   stn[9].wipBtn[48,0] := 0;
   stn[9].wipBtn[48,1] := 0;
   stn[9].wipBtn[48,2] := 0;
   stn[9].wipBtn[48,3] := 0;
   stn[9].wipBtn[48,4] := 0;
   stn[9].wipBtn[48,5] := 0;
   stn[9].wipBtn[48,6] := 0;
   stn[9].wipBtn[48,7] := 0;
   stn[9].wipBtn[49,0] := 0;
   stn[9].wipBtn[49,1] := 0;
   stn[9].wipBtn[49,2] := 0;
   stn[9].wipBtn[49,3] := 0;
   stn[9].wipBtn[49,4] := 0;
   stn[9].wipBtn[49,5] := 0;
   stn[9].wipBtn[49,6] := 0;
   stn[9].wipBtn[49,7] := 0;
   stn[10].wipBtn[0,0] := 0;
   stn[10].wipBtn[0,1] := 0;
   stn[10].wipBtn[0,2] := 0;
   stn[10].wipBtn[0,3] := 170;
   stn[10].wipBtn[0,4] := 0;
   stn[10].wipBtn[0,5] := 0;
   stn[10].wipBtn[1,0] := 0;
   stn[10].wipBtn[1,1] := 0;
   stn[10].wipBtn[1,2] := 0;
   stn[10].wipBtn[1,3] := 0;
   stn[10].wipBtn[1,4] := 0;
   stn[10].wipBtn[1,5] := 0;
   stn[10].wipBtn[1,6] := 0;
   stn[10].wipBtn[1,7] := 0;
   stn[10].wipBtn[2,0] := 0;
   stn[10].wipBtn[2,1] := 0;
   stn[10].wipBtn[2,2] := 0;
   stn[10].wipBtn[2,3] := 0;
   stn[10].wipBtn[2,4] := 0;
   stn[10].wipBtn[2,5] := 0;
   stn[10].wipBtn[2,6] := 0;
   stn[10].wipBtn[2,7] := 0;
   stn[10].wipBtn[3,0] := 0;
   stn[10].wipBtn[3,1] := 0;
   stn[10].wipBtn[3,2] := 0;
   stn[10].wipBtn[3,3] := 0;
   stn[10].wipBtn[3,4] := 0;
   stn[10].wipBtn[3,5] := 0;
   stn[10].wipBtn[3,6] := 0;
   stn[10].wipBtn[3,7] := 0;
   stn[10].wipBtn[4,0] := 0;
   stn[10].wipBtn[4,1] := 0;
   stn[10].wipBtn[4,2] := 0;
   stn[10].wipBtn[4,3] := 0;
   stn[10].wipBtn[4,4] := 0;
   stn[10].wipBtn[4,5] := 0;
   stn[10].wipBtn[4,6] := 0;
   stn[10].wipBtn[4,7] := 0;
   stn[10].wipBtn[5,0] := 0;
   stn[10].wipBtn[5,1] := 0;
   stn[10].wipBtn[5,2] := 0;
   stn[10].wipBtn[5,3] := 0;
   stn[10].wipBtn[5,4] := 0;
   stn[10].wipBtn[5,5] := 0;
   stn[10].wipBtn[5,6] := 0;
   stn[10].wipBtn[5,7] := 0;
   stn[10].wipBtn[6,0] := 0;
   stn[10].wipBtn[6,1] := 0;
   stn[10].wipBtn[6,2] := 0;
   stn[10].wipBtn[6,3] := 0;
   stn[10].wipBtn[6,4] := 0;
   stn[10].wipBtn[6,5] := 0;
   stn[10].wipBtn[6,6] := 0;
   stn[10].wipBtn[6,7] := 0;
   stn[10].wipBtn[7,0] := 0;
   stn[10].wipBtn[7,1] := 0;
   stn[10].wipBtn[7,2] := 0;
   stn[10].wipBtn[7,3] := 0;
   stn[10].wipBtn[7,4] := 0;
   stn[10].wipBtn[7,5] := 0;
   stn[10].wipBtn[7,6] := 0;
   stn[10].wipBtn[7,7] := 0;
   stn[10].wipBtn[8,0] := 0;
   stn[10].wipBtn[8,1] := 0;
   stn[10].wipBtn[8,2] := 0;
   stn[10].wipBtn[8,3] := 0;
   stn[10].wipBtn[8,4] := 0;
   stn[10].wipBtn[8,5] := 0;
   stn[10].wipBtn[8,6] := 0;
   stn[10].wipBtn[8,7] := 0;
   stn[10].wipBtn[9,0] := 0;
   stn[10].wipBtn[9,1] := 0;
   stn[10].wipBtn[9,2] := 0;
   stn[10].wipBtn[9,3] := 0;
   stn[10].wipBtn[9,4] := 0;
   stn[10].wipBtn[9,5] := 0;
   stn[10].wipBtn[9,6] := 0;
   stn[10].wipBtn[9,7] := 0;
   stn[10].wipBtn[10,0] := 0;
   stn[10].wipBtn[10,1] := 0;
   stn[10].wipBtn[10,2] := 0;
   stn[10].wipBtn[10,3] := 0;
   stn[10].wipBtn[10,4] := 0;
   stn[10].wipBtn[10,5] := 0;
   stn[10].wipBtn[10,6] := 0;
   stn[10].wipBtn[10,7] := 0;
   stn[10].wipBtn[11,0] := 0;
   stn[10].wipBtn[11,1] := 0;
   stn[10].wipBtn[11,2] := 0;
   stn[10].wipBtn[11,3] := 0;
   stn[10].wipBtn[11,4] := 0;
   stn[10].wipBtn[11,5] := 0;
   stn[10].wipBtn[11,6] := 0;
   stn[10].wipBtn[11,7] := 0;
   stn[10].wipBtn[12,0] := 0;
   stn[10].wipBtn[12,1] := 0;
   stn[10].wipBtn[12,2] := 0;
   stn[10].wipBtn[12,3] := 0;
   stn[10].wipBtn[12,4] := 0;
   stn[10].wipBtn[12,5] := 0;
   stn[10].wipBtn[12,6] := 0;
   stn[10].wipBtn[12,7] := 0;
   stn[10].wipBtn[13,0] := 0;
   stn[10].wipBtn[13,1] := 0;
   stn[10].wipBtn[13,2] := 0;
   stn[10].wipBtn[13,3] := 0;
   stn[10].wipBtn[13,4] := 0;
   stn[10].wipBtn[13,5] := 0;
   stn[10].wipBtn[13,6] := 0;
   stn[10].wipBtn[13,7] := 0;
   stn[10].wipBtn[14,0] := 0;
   stn[10].wipBtn[14,1] := 0;
   stn[10].wipBtn[14,2] := 0;
   stn[10].wipBtn[14,3] := 0;
   stn[10].wipBtn[14,4] := 0;
   stn[10].wipBtn[14,5] := 0;
   stn[10].wipBtn[14,6] := 0;
   stn[10].wipBtn[14,7] := 0;
   stn[10].wipBtn[15,0] := 0;
   stn[10].wipBtn[15,1] := 0;
   stn[10].wipBtn[15,2] := 0;
   stn[10].wipBtn[15,3] := 0;
   stn[10].wipBtn[15,4] := 0;
   stn[10].wipBtn[15,5] := 0;
   stn[10].wipBtn[15,6] := 0;
   stn[10].wipBtn[15,7] := 0;
   stn[10].wipBtn[16,0] := 0;
   stn[10].wipBtn[16,1] := 0;
   stn[10].wipBtn[16,2] := 0;
   stn[10].wipBtn[16,3] := 0;
   stn[10].wipBtn[16,4] := 0;
   stn[10].wipBtn[16,5] := 0;
   stn[10].wipBtn[16,6] := 0;
   stn[10].wipBtn[16,7] := 0;
   stn[10].wipBtn[17,0] := 0;
   stn[10].wipBtn[17,1] := 0;
   stn[10].wipBtn[17,2] := 0;
   stn[10].wipBtn[17,3] := 0;
   stn[10].wipBtn[17,4] := 0;
   stn[10].wipBtn[17,5] := 0;
   stn[10].wipBtn[17,6] := 0;
   stn[10].wipBtn[17,7] := 0;
   stn[10].wipBtn[18,0] := 0;
   stn[10].wipBtn[18,1] := 0;
   stn[10].wipBtn[18,2] := 0;
   stn[10].wipBtn[18,3] := 0;
   stn[10].wipBtn[18,4] := 0;
   stn[10].wipBtn[18,5] := 0;
   stn[10].wipBtn[18,6] := 0;
   stn[10].wipBtn[18,7] := 0;
   stn[10].wipBtn[19,0] := 0;
   stn[10].wipBtn[19,1] := 0;
   stn[10].wipBtn[19,2] := 0;
   stn[10].wipBtn[19,3] := 0;
   stn[10].wipBtn[19,4] := 0;
   stn[10].wipBtn[19,5] := 0;
   stn[10].wipBtn[19,6] := 0;
   stn[10].wipBtn[19,7] := 0;
   stn[10].wipBtn[20,0] := 0;
   stn[10].wipBtn[20,1] := 0;
   stn[10].wipBtn[20,2] := 0;
   stn[10].wipBtn[20,3] := 0;
   stn[10].wipBtn[20,4] := 0;
   stn[10].wipBtn[20,5] := 0;
   stn[10].wipBtn[20,6] := 0;
   stn[10].wipBtn[20,7] := 0;
   stn[10].wipBtn[21,0] := 0;
   stn[10].wipBtn[21,1] := 0;
   stn[10].wipBtn[21,2] := 0;
   stn[10].wipBtn[21,3] := 0;
   stn[10].wipBtn[21,4] := 0;
   stn[10].wipBtn[21,5] := 0;
   stn[10].wipBtn[21,6] := 0;
   stn[10].wipBtn[21,7] := 0;
   stn[10].wipBtn[22,0] := 0;
   stn[10].wipBtn[22,1] := 0;
   stn[10].wipBtn[22,2] := 0;
   stn[10].wipBtn[22,3] := 0;
   stn[10].wipBtn[22,4] := 0;
   stn[10].wipBtn[22,5] := 0;
   stn[10].wipBtn[22,6] := 0;
   stn[10].wipBtn[22,7] := 0;
   stn[10].wipBtn[23,0] := 0;
   stn[10].wipBtn[23,1] := 0;
   stn[10].wipBtn[23,2] := 0;
   stn[10].wipBtn[23,3] := 0;
   stn[10].wipBtn[23,4] := 0;
   stn[10].wipBtn[23,5] := 0;
   stn[10].wipBtn[23,6] := 0;
   stn[10].wipBtn[23,7] := 0;
   stn[10].wipBtn[24,0] := 0;
   stn[10].wipBtn[24,1] := 0;
   stn[10].wipBtn[24,2] := 0;
   stn[10].wipBtn[24,3] := 0;
   stn[10].wipBtn[24,4] := 0;
   stn[10].wipBtn[24,5] := 0;
   stn[10].wipBtn[24,6] := 0;
   stn[10].wipBtn[24,7] := 0;
   stn[10].wipBtn[25,0] := 0;
   stn[10].wipBtn[25,1] := 0;
   stn[10].wipBtn[25,2] := 0;
   stn[10].wipBtn[25,3] := 0;
   stn[10].wipBtn[25,4] := 0;
   stn[10].wipBtn[25,5] := 0;
   stn[10].wipBtn[25,6] := 0;
   stn[10].wipBtn[25,7] := 0;
   stn[10].wipBtn[26,0] := 0;
   stn[10].wipBtn[26,1] := 0;
   stn[10].wipBtn[26,2] := 0;
   stn[10].wipBtn[26,3] := 0;
   stn[10].wipBtn[26,4] := 0;
   stn[10].wipBtn[26,5] := 0;
   stn[10].wipBtn[26,6] := 0;
   stn[10].wipBtn[26,7] := 0;
   stn[10].wipBtn[27,0] := 0;
   stn[10].wipBtn[27,1] := 0;
   stn[10].wipBtn[27,2] := 0;
   stn[10].wipBtn[27,3] := 0;
   stn[10].wipBtn[27,4] := 0;
   stn[10].wipBtn[27,5] := 0;
   stn[10].wipBtn[27,6] := 0;
   stn[10].wipBtn[27,7] := 0;
   stn[10].wipBtn[28,0] := 0;
   stn[10].wipBtn[28,1] := 0;
   stn[10].wipBtn[28,2] := 0;
   stn[10].wipBtn[28,3] := 0;
   stn[10].wipBtn[28,4] := 0;
   stn[10].wipBtn[28,5] := 0;
   stn[10].wipBtn[28,6] := 0;
   stn[10].wipBtn[28,7] := 0;
   stn[10].wipBtn[29,0] := 0;
   stn[10].wipBtn[29,1] := 0;
   stn[10].wipBtn[29,2] := 0;
   stn[10].wipBtn[29,3] := 0;
   stn[10].wipBtn[29,4] := 0;
   stn[10].wipBtn[29,5] := 0;
   stn[10].wipBtn[29,6] := 0;
   stn[10].wipBtn[29,7] := 0;
   stn[10].wipBtn[30,0] := 0;
   stn[10].wipBtn[30,1] := 0;
   stn[10].wipBtn[30,2] := 0;
   stn[10].wipBtn[30,3] := 0;
   stn[10].wipBtn[30,4] := 0;
   stn[10].wipBtn[30,5] := 0;
   stn[10].wipBtn[30,6] := 0;
   stn[10].wipBtn[30,7] := 0;
   stn[10].wipBtn[31,0] := 0;
   stn[10].wipBtn[31,1] := 0;
   stn[10].wipBtn[31,2] := 0;
   stn[10].wipBtn[31,3] := 0;
   stn[10].wipBtn[31,4] := 0;
   stn[10].wipBtn[31,5] := 0;
   stn[10].wipBtn[31,6] := 0;
   stn[10].wipBtn[31,7] := 0;
   stn[10].wipBtn[32,0] := 0;
   stn[10].wipBtn[32,1] := 0;
   stn[10].wipBtn[32,2] := 0;
   stn[10].wipBtn[32,3] := 0;
   stn[10].wipBtn[32,4] := 0;
   stn[10].wipBtn[32,5] := 0;
   stn[10].wipBtn[32,6] := 0;
   stn[10].wipBtn[32,7] := 0;
   stn[10].wipBtn[33,0] := 0;
   stn[10].wipBtn[33,1] := 0;
   stn[10].wipBtn[33,2] := 0;
   stn[10].wipBtn[33,3] := 0;
   stn[10].wipBtn[33,4] := 0;
   stn[10].wipBtn[33,5] := 0;
   stn[10].wipBtn[33,6] := 0;
   stn[10].wipBtn[33,7] := 0;
   stn[10].wipBtn[34,0] := 0;
   stn[10].wipBtn[34,1] := 0;
   stn[10].wipBtn[34,2] := 0;
   stn[10].wipBtn[34,3] := 0;
   stn[10].wipBtn[34,4] := 0;
   stn[10].wipBtn[34,5] := 0;
   stn[10].wipBtn[34,6] := 0;
   stn[10].wipBtn[34,7] := 0;
   stn[10].wipBtn[35,0] := 0;
   stn[10].wipBtn[35,1] := 0;
   stn[10].wipBtn[35,2] := 0;
   stn[10].wipBtn[35,3] := 0;
   stn[10].wipBtn[35,4] := 0;
   stn[10].wipBtn[35,5] := 0;
   stn[10].wipBtn[35,6] := 0;
   stn[10].wipBtn[35,7] := 0;
   stn[10].wipBtn[36,0] := 0;
   stn[10].wipBtn[36,1] := 0;
   stn[10].wipBtn[36,2] := 0;
   stn[10].wipBtn[36,3] := 0;
   stn[10].wipBtn[36,4] := 0;
   stn[10].wipBtn[36,5] := 0;
   stn[10].wipBtn[36,6] := 0;
   stn[10].wipBtn[36,7] := 0;
   stn[10].wipBtn[37,0] := 0;
   stn[10].wipBtn[37,1] := 0;
   stn[10].wipBtn[37,2] := 0;
   stn[10].wipBtn[37,3] := 0;
   stn[10].wipBtn[37,4] := 0;
   stn[10].wipBtn[37,5] := 0;
   stn[10].wipBtn[37,6] := 0;
   stn[10].wipBtn[37,7] := 0;
   stn[10].wipBtn[38,0] := 0;
   stn[10].wipBtn[38,1] := 0;
   stn[10].wipBtn[38,2] := 0;
   stn[10].wipBtn[38,3] := 0;
   stn[10].wipBtn[38,4] := 0;
   stn[10].wipBtn[38,5] := 0;
   stn[10].wipBtn[38,6] := 0;
   stn[10].wipBtn[38,7] := 0;
   stn[10].wipBtn[39,0] := 0;
   stn[10].wipBtn[39,1] := 0;
   stn[10].wipBtn[39,2] := 0;
   stn[10].wipBtn[39,3] := 0;
   stn[10].wipBtn[39,4] := 0;
   stn[10].wipBtn[39,5] := 0;
   stn[10].wipBtn[39,6] := 0;
   stn[10].wipBtn[39,7] := 0;
   stn[10].wipBtn[40,0] := 0;
   stn[10].wipBtn[40,1] := 0;
   stn[10].wipBtn[40,2] := 0;
   stn[10].wipBtn[40,3] := 0;
   stn[10].wipBtn[40,4] := 0;
   stn[10].wipBtn[40,5] := 0;
   stn[10].wipBtn[40,6] := 0;
   stn[10].wipBtn[40,7] := 0;
   stn[10].wipBtn[41,0] := 0;
   stn[10].wipBtn[41,1] := 0;
   stn[10].wipBtn[41,2] := 0;
   stn[10].wipBtn[41,3] := 0;
   stn[10].wipBtn[41,4] := 0;
   stn[10].wipBtn[41,5] := 0;
   stn[10].wipBtn[41,6] := 0;
   stn[10].wipBtn[41,7] := 0;
   stn[10].wipBtn[42,0] := 0;
   stn[10].wipBtn[42,1] := 0;
   stn[10].wipBtn[42,2] := 0;
   stn[10].wipBtn[42,3] := 0;
   stn[10].wipBtn[42,4] := 0;
   stn[10].wipBtn[42,5] := 0;
   stn[10].wipBtn[42,6] := 0;
   stn[10].wipBtn[42,7] := 0;
   stn[10].wipBtn[43,0] := 0;
   stn[10].wipBtn[43,1] := 0;
   stn[10].wipBtn[43,2] := 0;
   stn[10].wipBtn[43,3] := 0;
   stn[10].wipBtn[43,4] := 0;
   stn[10].wipBtn[43,5] := 0;
   stn[10].wipBtn[43,6] := 0;
   stn[10].wipBtn[43,7] := 0;
   stn[10].wipBtn[44,0] := 0;
   stn[10].wipBtn[44,1] := 0;
   stn[10].wipBtn[44,2] := 0;
   stn[10].wipBtn[44,3] := 0;
   stn[10].wipBtn[44,4] := 0;
   stn[10].wipBtn[44,5] := 0;
   stn[10].wipBtn[44,6] := 0;
   stn[10].wipBtn[44,7] := 0;
   stn[10].wipBtn[45,0] := 0;
   stn[10].wipBtn[45,1] := 0;
   stn[10].wipBtn[45,2] := 0;
   stn[10].wipBtn[45,3] := 0;
   stn[10].wipBtn[45,4] := 0;
   stn[10].wipBtn[45,5] := 0;
   stn[10].wipBtn[45,6] := 0;
   stn[10].wipBtn[45,7] := 0;
   stn[10].wipBtn[46,0] := 0;
   stn[10].wipBtn[46,1] := 0;
   stn[10].wipBtn[46,2] := 0;
   stn[10].wipBtn[46,3] := 0;
   stn[10].wipBtn[46,4] := 0;
   stn[10].wipBtn[46,5] := 0;
   stn[10].wipBtn[46,6] := 0;
   stn[10].wipBtn[46,7] := 0;
   stn[10].wipBtn[47,0] := 0;
   stn[10].wipBtn[47,1] := 0;
   stn[10].wipBtn[47,2] := 0;
   stn[10].wipBtn[47,3] := 0;
   stn[10].wipBtn[47,4] := 0;
   stn[10].wipBtn[47,5] := 0;
   stn[10].wipBtn[47,6] := 0;
   stn[10].wipBtn[47,7] := 0;
   stn[10].wipBtn[48,0] := 0;
   stn[10].wipBtn[48,1] := 0;
   stn[10].wipBtn[48,2] := 0;
   stn[10].wipBtn[48,3] := 0;
   stn[10].wipBtn[48,4] := 0;
   stn[10].wipBtn[48,5] := 0;
   stn[10].wipBtn[48,6] := 0;
   stn[10].wipBtn[48,7] := 0;
   stn[10].wipBtn[49,0] := 0;
   stn[10].wipBtn[49,1] := 0;
   stn[10].wipBtn[49,2] := 0;
   stn[10].wipBtn[49,3] := 0;
   stn[10].wipBtn[49,4] := 0;
   stn[10].wipBtn[49,5] := 0;
   stn[10].wipBtn[49,6] := 0;
   stn[10].wipBtn[49,7] := 0;
   stn[11].wipBtn[0,0] := 0;
   stn[11].wipBtn[0,1] := 0;
   stn[11].wipBtn[0,2] := 0;
   stn[11].wipBtn[0,4] := 0;
   stn[11].wipBtn[0,5] := 0;
   stn[11].wipBtn[0,7] := 20;
   stn[11].wipBtn[1,0] := 0;
   stn[11].wipBtn[1,1] := 0;
   stn[11].wipBtn[1,2] := 0;
   stn[11].wipBtn[1,3] := 0;
   stn[11].wipBtn[1,4] := 0;
   stn[11].wipBtn[1,5] := 0;
   stn[11].wipBtn[1,6] := 0;
   stn[11].wipBtn[1,7] := 0;
   stn[11].wipBtn[2,0] := 0;
   stn[11].wipBtn[2,1] := 0;
   stn[11].wipBtn[2,2] := 0;
   stn[11].wipBtn[2,3] := 0;
   stn[11].wipBtn[2,4] := 0;
   stn[11].wipBtn[2,5] := 0;
   stn[11].wipBtn[2,6] := 0;
   stn[11].wipBtn[2,7] := 0;
   stn[11].wipBtn[3,0] := 0;
   stn[11].wipBtn[3,1] := 0;
   stn[11].wipBtn[3,2] := 0;
   stn[11].wipBtn[3,3] := 0;
   stn[11].wipBtn[3,4] := 0;
   stn[11].wipBtn[3,5] := 0;
   stn[11].wipBtn[3,6] := 0;
   stn[11].wipBtn[3,7] := 0;
   stn[11].wipBtn[4,0] := 0;
   stn[11].wipBtn[4,1] := 0;
   stn[11].wipBtn[4,2] := 0;
   stn[11].wipBtn[4,3] := 0;
   stn[11].wipBtn[4,4] := 0;
   stn[11].wipBtn[4,5] := 0;
   stn[11].wipBtn[4,6] := 0;
   stn[11].wipBtn[4,7] := 0;
   stn[11].wipBtn[5,0] := 0;
   stn[11].wipBtn[5,1] := 0;
   stn[11].wipBtn[5,2] := 0;
   stn[11].wipBtn[5,3] := 0;
   stn[11].wipBtn[5,4] := 0;
   stn[11].wipBtn[5,5] := 0;
   stn[11].wipBtn[5,6] := 0;
   stn[11].wipBtn[5,7] := 0;
   stn[11].wipBtn[6,0] := 0;
   stn[11].wipBtn[6,1] := 0;
   stn[11].wipBtn[6,2] := 0;
   stn[11].wipBtn[6,3] := 0;
   stn[11].wipBtn[6,4] := 0;
   stn[11].wipBtn[6,5] := 0;
   stn[11].wipBtn[6,6] := 0;
   stn[11].wipBtn[6,7] := 0;
   stn[11].wipBtn[7,0] := 0;
   stn[11].wipBtn[7,1] := 0;
   stn[11].wipBtn[7,2] := 0;
   stn[11].wipBtn[7,3] := 0;
   stn[11].wipBtn[7,4] := 0;
   stn[11].wipBtn[7,5] := 0;
   stn[11].wipBtn[7,6] := 0;
   stn[11].wipBtn[7,7] := 0;
   stn[11].wipBtn[8,0] := 0;
   stn[11].wipBtn[8,1] := 0;
   stn[11].wipBtn[8,2] := 0;
   stn[11].wipBtn[8,3] := 0;
   stn[11].wipBtn[8,4] := 0;
   stn[11].wipBtn[8,5] := 0;
   stn[11].wipBtn[8,6] := 0;
   stn[11].wipBtn[8,7] := 0;
   stn[11].wipBtn[9,0] := 0;
   stn[11].wipBtn[9,1] := 0;
   stn[11].wipBtn[9,2] := 0;
   stn[11].wipBtn[9,3] := 0;
   stn[11].wipBtn[9,4] := 0;
   stn[11].wipBtn[9,5] := 0;
   stn[11].wipBtn[9,6] := 0;
   stn[11].wipBtn[9,7] := 0;
   stn[11].wipBtn[10,0] := 0;
   stn[11].wipBtn[10,1] := 0;
   stn[11].wipBtn[10,2] := 0;
   stn[11].wipBtn[10,3] := 0;
   stn[11].wipBtn[10,4] := 0;
   stn[11].wipBtn[10,5] := 0;
   stn[11].wipBtn[10,6] := 0;
   stn[11].wipBtn[10,7] := 0;
   stn[11].wipBtn[11,0] := 0;
   stn[11].wipBtn[11,1] := 0;
   stn[11].wipBtn[11,2] := 0;
   stn[11].wipBtn[11,3] := 0;
   stn[11].wipBtn[11,4] := 0;
   stn[11].wipBtn[11,5] := 0;
   stn[11].wipBtn[11,6] := 0;
   stn[11].wipBtn[11,7] := 0;
   stn[11].wipBtn[12,0] := 0;
   stn[11].wipBtn[12,1] := 0;
   stn[11].wipBtn[12,2] := 0;
   stn[11].wipBtn[12,3] := 0;
   stn[11].wipBtn[12,4] := 0;
   stn[11].wipBtn[12,5] := 0;
   stn[11].wipBtn[12,6] := 0;
   stn[11].wipBtn[12,7] := 0;
   stn[11].wipBtn[13,0] := 0;
   stn[11].wipBtn[13,1] := 0;
   stn[11].wipBtn[13,2] := 0;
   stn[11].wipBtn[13,3] := 0;
   stn[11].wipBtn[13,4] := 0;
   stn[11].wipBtn[13,5] := 0;
   stn[11].wipBtn[13,6] := 0;
   stn[11].wipBtn[13,7] := 0;
   stn[11].wipBtn[14,0] := 0;
   stn[11].wipBtn[14,1] := 0;
   stn[11].wipBtn[14,2] := 0;
   stn[11].wipBtn[14,3] := 0;
   stn[11].wipBtn[14,4] := 0;
   stn[11].wipBtn[14,5] := 0;
   stn[11].wipBtn[14,6] := 0;
   stn[11].wipBtn[14,7] := 0;
   stn[11].wipBtn[15,0] := 0;
   stn[11].wipBtn[15,1] := 0;
   stn[11].wipBtn[15,2] := 0;
   stn[11].wipBtn[15,3] := 0;
   stn[11].wipBtn[15,4] := 0;
   stn[11].wipBtn[15,5] := 0;
   stn[11].wipBtn[15,6] := 0;
   stn[11].wipBtn[15,7] := 0;
   stn[11].wipBtn[16,0] := 0;
   stn[11].wipBtn[16,1] := 0;
   stn[11].wipBtn[16,2] := 0;
   stn[11].wipBtn[16,3] := 0;
   stn[11].wipBtn[16,4] := 0;
   stn[11].wipBtn[16,5] := 0;
   stn[11].wipBtn[16,6] := 0;
   stn[11].wipBtn[16,7] := 0;
   stn[11].wipBtn[17,0] := 0;
   stn[11].wipBtn[17,1] := 0;
   stn[11].wipBtn[17,2] := 0;
   stn[11].wipBtn[17,3] := 0;
   stn[11].wipBtn[17,4] := 0;
   stn[11].wipBtn[17,5] := 0;
   stn[11].wipBtn[17,6] := 0;
   stn[11].wipBtn[17,7] := 0;
   stn[11].wipBtn[18,0] := 0;
   stn[11].wipBtn[18,1] := 0;
   stn[11].wipBtn[18,2] := 0;
   stn[11].wipBtn[18,3] := 0;
   stn[11].wipBtn[18,4] := 0;
   stn[11].wipBtn[18,5] := 0;
   stn[11].wipBtn[18,6] := 0;
   stn[11].wipBtn[18,7] := 0;
   stn[11].wipBtn[19,0] := 0;
   stn[11].wipBtn[19,1] := 0;
   stn[11].wipBtn[19,2] := 0;
   stn[11].wipBtn[19,3] := 0;
   stn[11].wipBtn[19,4] := 0;
   stn[11].wipBtn[19,5] := 0;
   stn[11].wipBtn[19,6] := 0;
   stn[11].wipBtn[19,7] := 0;
   stn[11].wipBtn[20,0] := 0;
   stn[11].wipBtn[20,1] := 0;
   stn[11].wipBtn[20,2] := 0;
   stn[11].wipBtn[20,3] := 0;
   stn[11].wipBtn[20,4] := 0;
   stn[11].wipBtn[20,5] := 0;
   stn[11].wipBtn[20,6] := 0;
   stn[11].wipBtn[20,7] := 0;
   stn[11].wipBtn[21,0] := 0;
   stn[11].wipBtn[21,1] := 0;
   stn[11].wipBtn[21,2] := 0;
   stn[11].wipBtn[21,3] := 0;
   stn[11].wipBtn[21,4] := 0;
   stn[11].wipBtn[21,5] := 0;
   stn[11].wipBtn[21,6] := 0;
   stn[11].wipBtn[21,7] := 0;
   stn[11].wipBtn[22,0] := 0;
   stn[11].wipBtn[22,1] := 0;
   stn[11].wipBtn[22,2] := 0;
   stn[11].wipBtn[22,3] := 0;
   stn[11].wipBtn[22,4] := 0;
   stn[11].wipBtn[22,5] := 0;
   stn[11].wipBtn[22,6] := 0;
   stn[11].wipBtn[22,7] := 0;
   stn[11].wipBtn[23,0] := 0;
   stn[11].wipBtn[23,1] := 0;
   stn[11].wipBtn[23,2] := 0;
   stn[11].wipBtn[23,3] := 0;
   stn[11].wipBtn[23,4] := 0;
   stn[11].wipBtn[23,5] := 0;
   stn[11].wipBtn[23,6] := 0;
   stn[11].wipBtn[23,7] := 0;
   stn[11].wipBtn[24,0] := 0;
   stn[11].wipBtn[24,1] := 0;
   stn[11].wipBtn[24,2] := 0;
   stn[11].wipBtn[24,3] := 0;
   stn[11].wipBtn[24,4] := 0;
   stn[11].wipBtn[24,5] := 0;
   stn[11].wipBtn[24,6] := 0;
   stn[11].wipBtn[24,7] := 0;
   stn[11].wipBtn[25,0] := 0;
   stn[11].wipBtn[25,1] := 0;
   stn[11].wipBtn[25,2] := 0;
   stn[11].wipBtn[25,3] := 0;
   stn[11].wipBtn[25,4] := 0;
   stn[11].wipBtn[25,5] := 0;
   stn[11].wipBtn[25,6] := 0;
   stn[11].wipBtn[25,7] := 0;
   stn[11].wipBtn[26,0] := 0;
   stn[11].wipBtn[26,1] := 0;
   stn[11].wipBtn[26,2] := 0;
   stn[11].wipBtn[26,3] := 0;
   stn[11].wipBtn[26,4] := 0;
   stn[11].wipBtn[26,5] := 0;
   stn[11].wipBtn[26,6] := 0;
   stn[11].wipBtn[26,7] := 0;
   stn[11].wipBtn[27,0] := 0;
   stn[11].wipBtn[27,1] := 0;
   stn[11].wipBtn[27,2] := 0;
   stn[11].wipBtn[27,3] := 0;
   stn[11].wipBtn[27,4] := 0;
   stn[11].wipBtn[27,5] := 0;
   stn[11].wipBtn[27,6] := 0;
   stn[11].wipBtn[27,7] := 0;
   stn[11].wipBtn[28,0] := 0;
   stn[11].wipBtn[28,1] := 0;
   stn[11].wipBtn[28,2] := 0;
   stn[11].wipBtn[28,3] := 0;
   stn[11].wipBtn[28,4] := 0;
   stn[11].wipBtn[28,5] := 0;
   stn[11].wipBtn[28,6] := 0;
   stn[11].wipBtn[28,7] := 0;
   stn[11].wipBtn[29,0] := 0;
   stn[11].wipBtn[29,1] := 0;
   stn[11].wipBtn[29,2] := 0;
   stn[11].wipBtn[29,3] := 0;
   stn[11].wipBtn[29,4] := 0;
   stn[11].wipBtn[29,5] := 0;
   stn[11].wipBtn[29,6] := 0;
   stn[11].wipBtn[29,7] := 0;
   stn[11].wipBtn[30,0] := 0;
   stn[11].wipBtn[30,1] := 0;
   stn[11].wipBtn[30,2] := 0;
   stn[11].wipBtn[30,3] := 0;
   stn[11].wipBtn[30,4] := 0;
   stn[11].wipBtn[30,5] := 0;
   stn[11].wipBtn[30,6] := 0;
   stn[11].wipBtn[30,7] := 0;
   stn[11].wipBtn[31,0] := 0;
   stn[11].wipBtn[31,1] := 0;
   stn[11].wipBtn[31,2] := 0;
   stn[11].wipBtn[31,3] := 0;
   stn[11].wipBtn[31,4] := 0;
   stn[11].wipBtn[31,5] := 0;
   stn[11].wipBtn[31,6] := 0;
   stn[11].wipBtn[31,7] := 0;
   stn[11].wipBtn[32,0] := 0;
   stn[11].wipBtn[32,1] := 0;
   stn[11].wipBtn[32,2] := 0;
   stn[11].wipBtn[32,3] := 0;
   stn[11].wipBtn[32,4] := 0;
   stn[11].wipBtn[32,5] := 0;
   stn[11].wipBtn[32,6] := 0;
   stn[11].wipBtn[32,7] := 0;
   stn[11].wipBtn[33,0] := 0;
   stn[11].wipBtn[33,1] := 0;
   stn[11].wipBtn[33,2] := 0;
   stn[11].wipBtn[33,3] := 0;
   stn[11].wipBtn[33,4] := 0;
   stn[11].wipBtn[33,5] := 0;
   stn[11].wipBtn[33,6] := 0;
   stn[11].wipBtn[33,7] := 0;
   stn[11].wipBtn[34,0] := 0;
   stn[11].wipBtn[34,1] := 0;
   stn[11].wipBtn[34,2] := 0;
   stn[11].wipBtn[34,3] := 0;
   stn[11].wipBtn[34,4] := 0;
   stn[11].wipBtn[34,5] := 0;
   stn[11].wipBtn[34,6] := 0;
   stn[11].wipBtn[34,7] := 0;
   stn[11].wipBtn[35,0] := 0;
   stn[11].wipBtn[35,1] := 0;
   stn[11].wipBtn[35,2] := 0;
   stn[11].wipBtn[35,3] := 0;
   stn[11].wipBtn[35,4] := 0;
   stn[11].wipBtn[35,5] := 0;
   stn[11].wipBtn[35,6] := 0;
   stn[11].wipBtn[35,7] := 0;
   stn[11].wipBtn[36,0] := 0;
   stn[11].wipBtn[36,1] := 0;
   stn[11].wipBtn[36,2] := 0;
   stn[11].wipBtn[36,3] := 0;
   stn[11].wipBtn[36,4] := 0;
   stn[11].wipBtn[36,5] := 0;
   stn[11].wipBtn[36,6] := 0;
   stn[11].wipBtn[36,7] := 0;
   stn[11].wipBtn[37,0] := 0;
   stn[11].wipBtn[37,1] := 0;
   stn[11].wipBtn[37,2] := 0;
   stn[11].wipBtn[37,3] := 0;
   stn[11].wipBtn[37,4] := 0;
   stn[11].wipBtn[37,5] := 0;
   stn[11].wipBtn[37,6] := 0;
   stn[11].wipBtn[37,7] := 0;
   stn[11].wipBtn[38,0] := 0;
   stn[11].wipBtn[38,1] := 0;
   stn[11].wipBtn[38,2] := 0;
   stn[11].wipBtn[38,3] := 0;
   stn[11].wipBtn[38,4] := 0;
   stn[11].wipBtn[38,5] := 0;
   stn[11].wipBtn[38,6] := 0;
   stn[11].wipBtn[38,7] := 0;
   stn[11].wipBtn[39,0] := 0;
   stn[11].wipBtn[39,1] := 0;
   stn[11].wipBtn[39,2] := 0;
   stn[11].wipBtn[39,3] := 0;
   stn[11].wipBtn[39,4] := 0;
   stn[11].wipBtn[39,5] := 0;
   stn[11].wipBtn[39,6] := 0;
   stn[11].wipBtn[39,7] := 0;
   stn[11].wipBtn[40,0] := 0;
   stn[11].wipBtn[40,1] := 0;
   stn[11].wipBtn[40,2] := 0;
   stn[11].wipBtn[40,3] := 0;
   stn[11].wipBtn[40,4] := 0;
   stn[11].wipBtn[40,5] := 0;
   stn[11].wipBtn[40,6] := 0;
   stn[11].wipBtn[40,7] := 0;
   stn[11].wipBtn[41,0] := 0;
   stn[11].wipBtn[41,1] := 0;
   stn[11].wipBtn[41,2] := 0;
   stn[11].wipBtn[41,3] := 0;
   stn[11].wipBtn[41,4] := 0;
   stn[11].wipBtn[41,5] := 0;
   stn[11].wipBtn[41,6] := 0;
   stn[11].wipBtn[41,7] := 0;
   stn[11].wipBtn[42,0] := 0;
   stn[11].wipBtn[42,1] := 0;
   stn[11].wipBtn[42,2] := 0;
   stn[11].wipBtn[42,3] := 0;
   stn[11].wipBtn[42,4] := 0;
   stn[11].wipBtn[42,5] := 0;
   stn[11].wipBtn[42,6] := 0;
   stn[11].wipBtn[42,7] := 0;
   stn[11].wipBtn[43,0] := 0;
   stn[11].wipBtn[43,1] := 0;
   stn[11].wipBtn[43,2] := 0;
   stn[11].wipBtn[43,3] := 0;
   stn[11].wipBtn[43,4] := 0;
   stn[11].wipBtn[43,5] := 0;
   stn[11].wipBtn[43,6] := 0;
   stn[11].wipBtn[43,7] := 0;
   stn[11].wipBtn[44,0] := 0;
   stn[11].wipBtn[44,1] := 0;
   stn[11].wipBtn[44,2] := 0;
   stn[11].wipBtn[44,3] := 0;
   stn[11].wipBtn[44,4] := 0;
   stn[11].wipBtn[44,5] := 0;
   stn[11].wipBtn[44,6] := 0;
   stn[11].wipBtn[44,7] := 0;
   stn[11].wipBtn[45,0] := 0;
   stn[11].wipBtn[45,1] := 0;
   stn[11].wipBtn[45,2] := 0;
   stn[11].wipBtn[45,3] := 0;
   stn[11].wipBtn[45,4] := 0;
   stn[11].wipBtn[45,5] := 0;
   stn[11].wipBtn[45,6] := 0;
   stn[11].wipBtn[45,7] := 0;
   stn[11].wipBtn[46,0] := 0;
   stn[11].wipBtn[46,1] := 0;
   stn[11].wipBtn[46,2] := 0;
   stn[11].wipBtn[46,3] := 0;
   stn[11].wipBtn[46,4] := 0;
   stn[11].wipBtn[46,5] := 0;
   stn[11].wipBtn[46,6] := 0;
   stn[11].wipBtn[46,7] := 0;
   stn[11].wipBtn[47,0] := 0;
   stn[11].wipBtn[47,1] := 0;
   stn[11].wipBtn[47,2] := 0;
   stn[11].wipBtn[47,3] := 0;
   stn[11].wipBtn[47,4] := 0;
   stn[11].wipBtn[47,5] := 0;
   stn[11].wipBtn[47,6] := 0;
   stn[11].wipBtn[47,7] := 0;
   stn[11].wipBtn[48,0] := 0;
   stn[11].wipBtn[48,1] := 0;
   stn[11].wipBtn[48,2] := 0;
   stn[11].wipBtn[48,3] := 0;
   stn[11].wipBtn[48,4] := 0;
   stn[11].wipBtn[48,5] := 0;
   stn[11].wipBtn[48,6] := 0;
   stn[11].wipBtn[48,7] := 0;
   stn[11].wipBtn[49,0] := 0;
   stn[11].wipBtn[49,1] := 0;
   stn[11].wipBtn[49,2] := 0;
   stn[11].wipBtn[49,3] := 0;
   stn[11].wipBtn[49,4] := 0;
   stn[11].wipBtn[49,5] := 0;
   stn[11].wipBtn[49,6] := 0;
   stn[11].wipBtn[49,7] := 0;
   stn[12].wipBtn[0,0] := 0;
   stn[12].wipBtn[0,1] := 80;
   stn[12].wipBtn[0,4] := 0;
   stn[12].wipBtn[1,0] := 0;
   stn[12].wipBtn[1,1] := 0;
   stn[12].wipBtn[1,2] := 0;
   stn[12].wipBtn[1,3] := 0;
   stn[12].wipBtn[1,4] := 0;
   stn[12].wipBtn[1,5] := 0;
   stn[12].wipBtn[1,6] := 0;
   stn[12].wipBtn[1,7] := 0;
   stn[12].wipBtn[2,0] := 0;
   stn[12].wipBtn[2,1] := 0;
   stn[12].wipBtn[2,2] := 0;
   stn[12].wipBtn[2,3] := 0;
   stn[12].wipBtn[2,4] := 0;
   stn[12].wipBtn[2,5] := 0;
   stn[12].wipBtn[2,6] := 0;
   stn[12].wipBtn[2,7] := 0;
   stn[12].wipBtn[3,0] := 0;
   stn[12].wipBtn[3,1] := 0;
   stn[12].wipBtn[3,2] := 0;
   stn[12].wipBtn[3,3] := 0;
   stn[12].wipBtn[3,4] := 0;
   stn[12].wipBtn[3,5] := 0;
   stn[12].wipBtn[3,6] := 0;
   stn[12].wipBtn[3,7] := 0;
   stn[12].wipBtn[4,0] := 0;
   stn[12].wipBtn[4,1] := 0;
   stn[12].wipBtn[4,2] := 0;
   stn[12].wipBtn[4,3] := 0;
   stn[12].wipBtn[4,4] := 0;
   stn[12].wipBtn[4,5] := 0;
   stn[12].wipBtn[4,6] := 0;
   stn[12].wipBtn[4,7] := 0;
   stn[12].wipBtn[5,0] := 0;
   stn[12].wipBtn[5,1] := 0;
   stn[12].wipBtn[5,2] := 0;
   stn[12].wipBtn[5,3] := 0;
   stn[12].wipBtn[5,4] := 0;
   stn[12].wipBtn[5,5] := 0;
   stn[12].wipBtn[5,6] := 0;
   stn[12].wipBtn[5,7] := 0;
   stn[12].wipBtn[6,0] := 0;
   stn[12].wipBtn[6,1] := 0;
   stn[12].wipBtn[6,2] := 0;
   stn[12].wipBtn[6,3] := 0;
   stn[12].wipBtn[6,4] := 0;
   stn[12].wipBtn[6,5] := 0;
   stn[12].wipBtn[6,6] := 0;
   stn[12].wipBtn[6,7] := 0;
   stn[12].wipBtn[7,0] := 0;
   stn[12].wipBtn[7,1] := 0;
   stn[12].wipBtn[7,2] := 0;
   stn[12].wipBtn[7,3] := 0;
   stn[12].wipBtn[7,4] := 0;
   stn[12].wipBtn[7,5] := 0;
   stn[12].wipBtn[7,6] := 0;
   stn[12].wipBtn[7,7] := 0;
   stn[12].wipBtn[8,0] := 0;
   stn[12].wipBtn[8,1] := 0;
   stn[12].wipBtn[8,2] := 0;
   stn[12].wipBtn[8,3] := 0;
   stn[12].wipBtn[8,4] := 0;
   stn[12].wipBtn[8,5] := 0;
   stn[12].wipBtn[8,6] := 0;
   stn[12].wipBtn[8,7] := 0;
   stn[12].wipBtn[9,0] := 0;
   stn[12].wipBtn[9,1] := 0;
   stn[12].wipBtn[9,2] := 0;
   stn[12].wipBtn[9,3] := 0;
   stn[12].wipBtn[9,4] := 0;
   stn[12].wipBtn[9,5] := 0;
   stn[12].wipBtn[9,6] := 0;
   stn[12].wipBtn[9,7] := 0;
   stn[12].wipBtn[10,0] := 0;
   stn[12].wipBtn[10,1] := 0;
   stn[12].wipBtn[10,2] := 0;
   stn[12].wipBtn[10,3] := 0;
   stn[12].wipBtn[10,4] := 0;
   stn[12].wipBtn[10,5] := 0;
   stn[12].wipBtn[10,6] := 0;
   stn[12].wipBtn[10,7] := 0;
   stn[12].wipBtn[11,0] := 0;
   stn[12].wipBtn[11,1] := 0;
   stn[12].wipBtn[11,2] := 0;
   stn[12].wipBtn[11,3] := 0;
   stn[12].wipBtn[11,4] := 0;
   stn[12].wipBtn[11,5] := 0;
   stn[12].wipBtn[11,6] := 0;
   stn[12].wipBtn[11,7] := 0;
   stn[12].wipBtn[12,0] := 0;
   stn[12].wipBtn[12,1] := 0;
   stn[12].wipBtn[12,2] := 0;
   stn[12].wipBtn[12,3] := 0;
   stn[12].wipBtn[12,4] := 0;
   stn[12].wipBtn[12,5] := 0;
   stn[12].wipBtn[12,6] := 0;
   stn[12].wipBtn[12,7] := 0;
   stn[12].wipBtn[13,0] := 0;
   stn[12].wipBtn[13,1] := 0;
   stn[12].wipBtn[13,2] := 0;
   stn[12].wipBtn[13,3] := 0;
   stn[12].wipBtn[13,4] := 0;
   stn[12].wipBtn[13,5] := 0;
   stn[12].wipBtn[13,6] := 0;
   stn[12].wipBtn[13,7] := 0;
   stn[12].wipBtn[14,0] := 0;
   stn[12].wipBtn[14,1] := 0;
   stn[12].wipBtn[14,2] := 0;
   stn[12].wipBtn[14,3] := 0;
   stn[12].wipBtn[14,4] := 0;
   stn[12].wipBtn[14,5] := 0;
   stn[12].wipBtn[14,6] := 0;
   stn[12].wipBtn[14,7] := 0;
   stn[12].wipBtn[15,0] := 0;
   stn[12].wipBtn[15,1] := 0;
   stn[12].wipBtn[15,2] := 0;
   stn[12].wipBtn[15,3] := 0;
   stn[12].wipBtn[15,4] := 0;
   stn[12].wipBtn[15,5] := 0;
   stn[12].wipBtn[15,6] := 0;
   stn[12].wipBtn[15,7] := 0;
   stn[12].wipBtn[16,0] := 0;
   stn[12].wipBtn[16,1] := 0;
   stn[12].wipBtn[16,2] := 0;
   stn[12].wipBtn[16,3] := 0;
   stn[12].wipBtn[16,4] := 0;
   stn[12].wipBtn[16,5] := 0;
   stn[12].wipBtn[16,6] := 0;
   stn[12].wipBtn[16,7] := 0;
   stn[12].wipBtn[17,0] := 0;
   stn[12].wipBtn[17,1] := 0;
   stn[12].wipBtn[17,2] := 0;
   stn[12].wipBtn[17,3] := 0;
   stn[12].wipBtn[17,4] := 0;
   stn[12].wipBtn[17,5] := 0;
   stn[12].wipBtn[17,6] := 0;
   stn[12].wipBtn[17,7] := 0;
   stn[12].wipBtn[18,0] := 0;
   stn[12].wipBtn[18,1] := 0;
   stn[12].wipBtn[18,2] := 0;
   stn[12].wipBtn[18,3] := 0;
   stn[12].wipBtn[18,4] := 0;
   stn[12].wipBtn[18,5] := 0;
   stn[12].wipBtn[18,6] := 0;
   stn[12].wipBtn[18,7] := 0;
   stn[12].wipBtn[19,0] := 0;
   stn[12].wipBtn[19,1] := 0;
   stn[12].wipBtn[19,2] := 0;
   stn[12].wipBtn[19,3] := 0;
   stn[12].wipBtn[19,4] := 0;
   stn[12].wipBtn[19,5] := 0;
   stn[12].wipBtn[19,6] := 0;
   stn[12].wipBtn[19,7] := 0;
   stn[12].wipBtn[20,0] := 0;
   stn[12].wipBtn[20,1] := 0;
   stn[12].wipBtn[20,2] := 0;
   stn[12].wipBtn[20,3] := 0;
   stn[12].wipBtn[20,4] := 0;
   stn[12].wipBtn[20,5] := 0;
   stn[12].wipBtn[20,6] := 0;
   stn[12].wipBtn[20,7] := 0;
   stn[12].wipBtn[21,0] := 0;
   stn[12].wipBtn[21,1] := 0;
   stn[12].wipBtn[21,2] := 0;
   stn[12].wipBtn[21,3] := 0;
   stn[12].wipBtn[21,4] := 0;
   stn[12].wipBtn[21,5] := 0;
   stn[12].wipBtn[21,6] := 0;
   stn[12].wipBtn[21,7] := 0;
   stn[12].wipBtn[22,0] := 0;
   stn[12].wipBtn[22,1] := 0;
   stn[12].wipBtn[22,2] := 0;
   stn[12].wipBtn[22,3] := 0;
   stn[12].wipBtn[22,4] := 0;
   stn[12].wipBtn[22,5] := 0;
   stn[12].wipBtn[22,6] := 0;
   stn[12].wipBtn[22,7] := 0;
   stn[12].wipBtn[23,0] := 0;
   stn[12].wipBtn[23,1] := 0;
   stn[12].wipBtn[23,2] := 0;
   stn[12].wipBtn[23,3] := 0;
   stn[12].wipBtn[23,4] := 0;
   stn[12].wipBtn[23,5] := 0;
   stn[12].wipBtn[23,6] := 0;
   stn[12].wipBtn[23,7] := 0;
   stn[12].wipBtn[24,0] := 0;
   stn[12].wipBtn[24,1] := 0;
   stn[12].wipBtn[24,2] := 0;
   stn[12].wipBtn[24,3] := 0;
   stn[12].wipBtn[24,4] := 0;
   stn[12].wipBtn[24,5] := 0;
   stn[12].wipBtn[24,6] := 0;
   stn[12].wipBtn[24,7] := 0;
   stn[12].wipBtn[25,0] := 0;
   stn[12].wipBtn[25,1] := 0;
   stn[12].wipBtn[25,2] := 0;
   stn[12].wipBtn[25,3] := 0;
   stn[12].wipBtn[25,4] := 0;
   stn[12].wipBtn[25,5] := 0;
   stn[12].wipBtn[25,6] := 0;
   stn[12].wipBtn[25,7] := 0;
   stn[12].wipBtn[26,0] := 0;
   stn[12].wipBtn[26,1] := 0;
   stn[12].wipBtn[26,2] := 0;
   stn[12].wipBtn[26,3] := 0;
   stn[12].wipBtn[26,4] := 0;
   stn[12].wipBtn[26,5] := 0;
   stn[12].wipBtn[26,6] := 0;
   stn[12].wipBtn[26,7] := 0;
   stn[12].wipBtn[27,0] := 0;
   stn[12].wipBtn[27,1] := 0;
   stn[12].wipBtn[27,2] := 0;
   stn[12].wipBtn[27,3] := 0;
   stn[12].wipBtn[27,4] := 0;
   stn[12].wipBtn[27,5] := 0;
   stn[12].wipBtn[27,6] := 0;
   stn[12].wipBtn[27,7] := 0;
   stn[12].wipBtn[28,0] := 0;
   stn[12].wipBtn[28,1] := 0;
   stn[12].wipBtn[28,2] := 0;
   stn[12].wipBtn[28,3] := 0;
   stn[12].wipBtn[28,4] := 0;
   stn[12].wipBtn[28,5] := 0;
   stn[12].wipBtn[28,6] := 0;
   stn[12].wipBtn[28,7] := 0;
   stn[12].wipBtn[29,0] := 0;
   stn[12].wipBtn[29,1] := 0;
   stn[12].wipBtn[29,2] := 0;
   stn[12].wipBtn[29,3] := 0;
   stn[12].wipBtn[29,4] := 0;
   stn[12].wipBtn[29,5] := 0;
   stn[12].wipBtn[29,6] := 0;
   stn[12].wipBtn[29,7] := 0;
   stn[12].wipBtn[30,0] := 0;
   stn[12].wipBtn[30,1] := 0;
   stn[12].wipBtn[30,2] := 0;
   stn[12].wipBtn[30,3] := 0;
   stn[12].wipBtn[30,4] := 0;
   stn[12].wipBtn[30,5] := 0;
   stn[12].wipBtn[30,6] := 0;
   stn[12].wipBtn[30,7] := 0;
   stn[12].wipBtn[31,0] := 0;
   stn[12].wipBtn[31,1] := 0;
   stn[12].wipBtn[31,2] := 0;
   stn[12].wipBtn[31,3] := 0;
   stn[12].wipBtn[31,4] := 0;
   stn[12].wipBtn[31,5] := 0;
   stn[12].wipBtn[31,6] := 0;
   stn[12].wipBtn[31,7] := 0;
   stn[12].wipBtn[32,0] := 0;
   stn[12].wipBtn[32,1] := 0;
   stn[12].wipBtn[32,2] := 0;
   stn[12].wipBtn[32,3] := 0;
   stn[12].wipBtn[32,4] := 0;
   stn[12].wipBtn[32,5] := 0;
   stn[12].wipBtn[32,6] := 0;
   stn[12].wipBtn[32,7] := 0;
   stn[12].wipBtn[33,0] := 0;
   stn[12].wipBtn[33,1] := 0;
   stn[12].wipBtn[33,2] := 0;
   stn[12].wipBtn[33,3] := 0;
   stn[12].wipBtn[33,4] := 0;
   stn[12].wipBtn[33,5] := 0;
   stn[12].wipBtn[33,6] := 0;
   stn[12].wipBtn[33,7] := 0;
   stn[12].wipBtn[34,0] := 0;
   stn[12].wipBtn[34,1] := 0;
   stn[12].wipBtn[34,2] := 0;
   stn[12].wipBtn[34,3] := 0;
   stn[12].wipBtn[34,4] := 0;
   stn[12].wipBtn[34,5] := 0;
   stn[12].wipBtn[34,6] := 0;
   stn[12].wipBtn[34,7] := 0;
   stn[12].wipBtn[35,0] := 0;
   stn[12].wipBtn[35,1] := 0;
   stn[12].wipBtn[35,2] := 0;
   stn[12].wipBtn[35,3] := 0;
   stn[12].wipBtn[35,4] := 0;
   stn[12].wipBtn[35,5] := 0;
   stn[12].wipBtn[35,6] := 0;
   stn[12].wipBtn[35,7] := 0;
   stn[12].wipBtn[36,0] := 0;
   stn[12].wipBtn[36,1] := 0;
   stn[12].wipBtn[36,2] := 0;
   stn[12].wipBtn[36,3] := 0;
   stn[12].wipBtn[36,4] := 0;
   stn[12].wipBtn[36,5] := 0;
   stn[12].wipBtn[36,6] := 0;
   stn[12].wipBtn[36,7] := 0;
   stn[12].wipBtn[37,0] := 0;
   stn[12].wipBtn[37,1] := 0;
   stn[12].wipBtn[37,2] := 0;
   stn[12].wipBtn[37,3] := 0;
   stn[12].wipBtn[37,4] := 0;
   stn[12].wipBtn[37,5] := 0;
   stn[12].wipBtn[37,6] := 0;
   stn[12].wipBtn[37,7] := 0;
   stn[12].wipBtn[38,0] := 0;
   stn[12].wipBtn[38,1] := 0;
   stn[12].wipBtn[38,2] := 0;
   stn[12].wipBtn[38,3] := 0;
   stn[12].wipBtn[38,4] := 0;
   stn[12].wipBtn[38,5] := 0;
   stn[12].wipBtn[38,6] := 0;
   stn[12].wipBtn[38,7] := 0;